// Mitsubishi GX Works2 project: 70常温静置库1130   PLC: Q10UDEH (continued)
		m_iCoordinateY:=1;
		FanucRobotIO.io_xMutexLock:=0;
	END_IF;
	IF ConveyorIO.xEmpty AND PackCommunicationIO.o_iSinglePackDonePLCPC=1 THEN
		m_iStep:=1;
	END_IF;
END_CASE;
END_FUNCTION_BLOCK

PROGRAM POU
VAR
  Conveyor70101 : Conveyor;
  Conveyor70102 : Conveyor;
  Conveyor70103 : Conveyor;
  Conveyor70104 : Conveyor;
  Conveyor70105 : Conveyor;
  Conveyor70106 : Conveyor;
  Conveyor70107 : Conveyor;
  Conveyor70108 : Conveyor;
  Conveyor70109 : Conveyor;
  Conveyor70110 : Conveyor;
  Conveyor70111 : Conveyor;
  Conveyor70112 : Conveyor;
  Conveyor70113 : Conveyor;
  Conveyor70114 : Conveyor;
  Conveyor70115 : Conveyor;
  Conveyor70116 : Conveyor;
  Conveyor70117 : Conveyor;
  Conveyor70118 : Conveyor;
  Conveyor70119 : Conveyor;
  Conveyor70120 : Conveyor;
  Conveyor70121 : Conveyor;
  Conveyor70122 : Conveyor;
  Conveyor70123 : Conveyor;
  Conveyor70124 : Conveyor;
  Conveyor70125 : Conveyor;
  Conveyor70126 : Conveyor;
  Conveyor70127 : Conveyor;
  Conveyor70128 : Conveyor;
  Conveyor70129 : Conveyor;
  Conveyor70130 : Conveyor;
  Conveyor70131 : Conveyor;
  Conveyor70132 : Conveyor;
  Conveyor70133 : Conveyor;
  Conveyor70134 : Conveyor;
  Conveyor70135 : Conveyor;
  Conveyor70136 : Conveyor;
  Conveyor70137 : Conveyor;
  Conveyor70138 : Conveyor;
  Conveyor70139 : Conveyor;
  Conveyor70140 : Conveyor;
  Conveyor70141 : Conveyor;
  Conveyor70142 : Conveyor;
  Conveyor70143 : Conveyor;
  Conveyor70144 : Conveyor;
  Conveyor70145 : Conveyor;
  Conveyor70146 : Conveyor;
  Conveyor70147 : Conveyor;
  Conveyor70148 : Conveyor;
  Conveyor70149 : Conveyor;
  Conveyor70150 : Conveyor;
  Conveyor70151 : Conveyor;
  Conveyor70152 : Conveyor;
  Conveyor70153 : Conveyor;
  Conveyor70154 : Conveyor;
  Conveyor70155 : Conveyor;
  Conveyor70156 : Conveyor;
  Conveyor70157 : Conveyor;
  Conveyor70158 : Conveyor;
  Conveyor70159 : Conveyor;
  Conveyor70160 : Conveyor;
  Conveyor70161 : Conveyor;
  Conveyor70162 : Conveyor;
  Conveyor70163 : Conveyor;
  Conveyor70164 : Conveyor;
  Conveyor70165 : Conveyor;
  Conveyor70166 : Conveyor;
  Conveyor70167 : Conveyor;
  Conveyor70168 : Conveyor;
  Conveyor70169 : Conveyor;
  Conveyor70170 : Conveyor;
  Conveyor70171 : Conveyor;
  Conveyor70172 : Conveyor;
  Conveyor70173 : Conveyor;
  Conveyor70174 : Conveyor;
  Conveyor70175 : Conveyor;
  Conveyor70176 : Conveyor;
  Conveyor70177 : Conveyor;
  Conveyor70178 : Conveyor;
  Conveyor70179 : Conveyor;
  Conveyor70180 : Conveyor;
  Conveyor70181 : Conveyor;
  Conveyor70182 : Conveyor;
  Conveyor70183 : Conveyor;
  Conveyor70184 : Conveyor;
  Conveyor70185 : Conveyor;
  Conveyor70186 : Conveyor;
  Conveyor70187 : Conveyor;
  Conveyor70188 : Conveyor;
  Conveyor70189 : Conveyor;
  Conveyor70190 : Conveyor;
  Conveyor70191 : Conveyor;
  Conveyor70192 : Conveyor;
  Conveyor70193 : Conveyor;
  Conveyor70194 : Conveyor;
  Conveyor70195 : Conveyor;
  Conveyor70196 : Conveyor;
  Conveyor70197 : Conveyor;
  Conveyor70198 : Conveyor;
  Conveyor70199 : Conveyor;
  Conveyor701100 : Conveyor;
  Conveyor701101 : Conveyor;
  Conveyor701102 : Conveyor;
  Conveyor701103 : Conveyor;
  Conveyor701104 : Conveyor;
  Conveyor701105 : Conveyor;
  Conveyor701106 : Conveyor;
  Conveyor701107 : Conveyor;
  Conveyor701108 : Conveyor;
  Conveyor701109 : Conveyor;
  Conveyor701110 : Conveyor;
  Conveyor701111 : Conveyor;
  Conveyor701112 : Conveyor;
  ConveyorIO70101 : ConveyorIO;
  ConveyorIO70102 : ConveyorIO;
  ConveyorIO70103 : ConveyorIO;
  ConveyorIO70104 : ConveyorIO;
  ConveyorIO70105 : ConveyorIO;
  ConveyorIO70106 : ConveyorIO;
  ConveyorIO70107 : ConveyorIO;
  ConveyorIO70108 : ConveyorIO;
  ConveyorIO70109 : ConveyorIO;
  ConveyorIO70110 : ConveyorIO;
  ConveyorIO70111 : ConveyorIO;
  ConveyorIO70112 : ConveyorIO;
  ConveyorIO70113 : ConveyorIO;
  ConveyorIO70114 : ConveyorIO;
  ConveyorIO70115 : ConveyorIO;
  ConveyorIO70116 : ConveyorIO;
  ConveyorIO70117 : ConveyorIO;
  ConveyorIO70118 : ConveyorIO;
  ConveyorIO70119 : ConveyorIO;
  ConveyorIO70120 : ConveyorIO;
  ConveyorIO70121 : ConveyorIO;
  ConveyorIO70122 : ConveyorIO;
  ConveyorIO70123 : ConveyorIO;
  ConveyorIO70124 : ConveyorIO;
  ConveyorIO70125 : ConveyorIO;
  ConveyorIO70126 : ConveyorIO;
  ConveyorIO70127 : ConveyorIO;
  ConveyorIO70128 : ConveyorIO;
  ConveyorIO70129 : ConveyorIO;
  ConveyorIO70130 : ConveyorIO;
  ConveyorIO70131 : ConveyorIO;
  ConveyorIO70132 : ConveyorIO;
  ConveyorIO70133 : ConveyorIO;
  ConveyorIO70134 : ConveyorIO;
  ConveyorIO70135 : ConveyorIO;
  ConveyorIO70136 : ConveyorIO;
  ConveyorIO70137 : ConveyorIO;
  ConveyorIO70138 : ConveyorIO;
  ConveyorIO70139 : ConveyorIO;
  ConveyorIO70140 : ConveyorIO;
  ConveyorIO70141 : ConveyorIO;
  ConveyorIO70142 : ConveyorIO;
  ConveyorIO70143 : ConveyorIO;
  ConveyorIO70144 : ConveyorIO;
  ConveyorIO70145 : ConveyorIO;
  ConveyorIO70146 : ConveyorIO;
  ConveyorIO70147 : ConveyorIO;
  ConveyorIO70148 : ConveyorIO;
  ConveyorIO70149 : ConveyorIO;
  ConveyorIO70150 : ConveyorIO;
  ConveyorIO70151 : ConveyorIO;
  ConveyorIO70152 : ConveyorIO;
  ConveyorIO70153 : ConveyorIO;
  ConveyorIO70154 : ConveyorIO;
  ConveyorIO70155 : ConveyorIO;
  ConveyorIO70156 : ConveyorIO;
  ConveyorIO70157 : ConveyorIO;
  ConveyorIO70158 : ConveyorIO;
  ConveyorIO70159 : ConveyorIO;
  ConveyorIO70160 : ConveyorIO;
  ConveyorIO70161 : ConveyorIO;
  ConveyorIO70162 : ConveyorIO;
  ConveyorIO70163 : ConveyorIO;
  ConveyorIO70164 : ConveyorIO;
  ConveyorIO70165 : ConveyorIO;
  ConveyorIO70166 : ConveyorIO;
  ConveyorIO70167 : ConveyorIO;
  ConveyorIO70168 : ConveyorIO;
  ConveyorIO70169 : ConveyorIO;
  ConveyorIO70170 : ConveyorIO;
  ConveyorIO70171 : ConveyorIO;
  ConveyorIO70172 : ConveyorIO;
  ConveyorIO70173 : ConveyorIO;
  ConveyorIO70174 : ConveyorIO;
  ConveyorIO70175 : ConveyorIO;
  ConveyorIO70176 : ConveyorIO;
  ConveyorIO70177 : ConveyorIO;
  ConveyorIO70178 : ConveyorIO;
  ConveyorIO70179 : ConveyorIO;
  ConveyorIO70180 : ConveyorIO;
  ConveyorIO70181 : ConveyorIO;
  ConveyorIO70182 : ConveyorIO;
  ConveyorIO70183 : ConveyorIO;
  ConveyorIO70184 : ConveyorIO;
  ConveyorIO70185 : ConveyorIO;
  ConveyorIO70186 : ConveyorIO;
  ConveyorIO70187 : ConveyorIO;
  ConveyorIO70188 : ConveyorIO;
  ConveyorIO70189 : ConveyorIO;
  ConveyorIO70190 : ConveyorIO;
  ConveyorIO70191 : ConveyorIO;
  ConveyorIO70192 : ConveyorIO;
  ConveyorIO70193 : ConveyorIO;
  ConveyorIO70194 : ConveyorIO;
  ConveyorIO70195 : ConveyorIO;
  ConveyorIO70196 : ConveyorIO;
  ConveyorIO70197 : ConveyorIO;
  ConveyorIO70198 : ConveyorIO;
  ConveyorIO70199 : ConveyorIO;
  ConveyorIO701100 : ConveyorIO;
  ConveyorIO701101 : ConveyorIO;
  ConveyorIO701102 : ConveyorIO;
  ConveyorIO701103 : ConveyorIO;
  ConveyorIO701104 : ConveyorIO;
  ConveyorIO701105 : ConveyorIO;
  ConveyorIO701106 : ConveyorIO;
  ConveyorIO701107 : ConveyorIO;
  ConveyorIO701108 : ConveyorIO;
  ConveyorIO701109 : ConveyorIO;
  ConveyorIO701110 : ConveyorIO;
  ConveyorIO701111 : ConveyorIO;
  ConveyorIO701112 : ConveyorIO;
  Switch70301 : Switch;
  SwitchIO70301 : SwitchIO;
  Lift70207 : ShuttleCar;
  LifterIO70207 : ShuttleCarIO;
  ConveyorIO701113 : ConveyorIO;
  ConveyorIO701114 : ConveyorIO;
  ConveyorIO701115 : ConveyorIO;
  ConveyorIO701116 : ConveyorIO;
  ConveyorIO701117 : ConveyorIO;
  ConveyorIO701118 : ConveyorIO;
  ConveyorIO701119 : ConveyorIO;
  ConveyorIO701120 : ConveyorIO;
  Conveyor701113 : Conveyor;
  Conveyor701114 : Conveyor;
  Conveyor701115 : Conveyor;
  Conveyor701116 : Conveyor;
  Conveyor701117 : Conveyor;
  Conveyor701118 : Conveyor;
  Conveyor701119 : Conveyor;
  Conveyor701120 : Conveyor;
  Switch70326 : Switch;
  SwitchIO70326 : SwitchIO;
  Conveyor701111_1 : Conveyor;
  ConveyorIO701111_1 : ConveyorIO;
  Switch70311 : Switch;
  SwitchIO70311 : SwitchIO;
  Switch70316 : Switch;
  SwitchIO70316 : SwitchIO;
  m_xRGVSemiAuto : BOOL;
  m_iRGVDestinationPos : INT;
  m_xRGVReset : BOOL;
  m_iRGVCurrentPos : INT;
  m_xRGVPositionArrive : BOOL;
  m_xRGVConveyorEmpty : BOOL;
  m_xRGVConveyorNextRun : BOOL;
  m_xRGVAlarm : BOOL;
  m_xtonConveyor70195Reset : TON;
  m_xtonConveyor70195CurTime : TIME;
  m_xtonConveyor70146Reset : TON;
  m_xtonConveyor70146CurTime : TIME;
  m_xtonConveyor701115Reset : TON;
  m_xtonConveyor701114Reset : TON;
  m_xtonConveyor701115CurTime : TIME;
  m_xtonConveyor701114CurTime : TIME;
  Switch70317 : Switch;
  SwitchIO70317 : SwitchIO;
  ConveyorIO70165_1 : ConveyorIO;
  Conveyor70165_1 : Conveyor;
  m_xOCV2_1LoadRequest : BOOL;  (* OCV2  1号机上料请求 *)
  m_xOCV2_1LoadStart : BOOL;  (* OCV2 1号机开始上料信号 *)
  m_xOCV2_1UnloadRequest : BOOL;  (* OCV2 1号机开始下料信号 *)
  m_xOCV2_2UnloadRequest : BOOL;  (* OCV2 2号机开始下料信号 *)
  Switch70318 : Switch;
  m_xOCV2_1UnloadStart : BOOL;  (* 允许下料 *)
  Switch70319 : Switch;
  SwitchIO70319 : SwitchIO;
  Switch70320 : Switch;
  SwitchIO70320 : SwitchIO;
  m_x60LoadRequest : BOOL;
  m_xOCV2_1LoadLock : BOOL;  (* OCV2上料自锁 *)
  m_xOCV2_1UnLoadLock : BOOL;  (* OCV2下料自锁 *)
  m_xOCV3_1LoadRequest : BOOL;  (* OCV3  1号机上料请求 *)
  m_xOCV3_1LoadStart : BOOL;  (* OCV3 1号机开始上料信号 *)
  m_xOCV3_1UnloadRequest : BOOL;  (* OCV3 1号机开始下料信号 *)
  m_xOCV3_1UnloadStart : BOOL;  (* OCV3  1号机下料请求 *)
  m_xOCV3_1LoadLock : BOOL;  (* OCV3——1上料自锁 *)
  m_xOCV3_1UnLoadLock : BOOL;  (* OCV3——1下料自锁 *)
  ConveyorIO70175_1 : ConveyorIO;
  Conveyor70175_1 : Conveyor;
  m_xtonConveyor70162Reset : TON;
  m_xtonConveyor70162CurTime : TIME;
  m_xtonConveyor701103Reset : TON;
  m_xtonConveyor701103CurTime : TIME;
  m_xtonConveyor70159Reset : TON;
  m_xtonConveyor70159CurTime : TIME;
  m_xtonConveyor701102Reset : TON;
  m_xtonConveyor701102CurTime : TIME;
  m_xtonConveyor70170Reset : TON;
  m_xtonConveyor70170CurTime : TIME;
  m_xtonConveyor70168Reset : TON;
  m_xtonConveyor70168CurTime : TIME;
  m_xOCV2_2LoadRequest : BOOL;  (* OCV2 2号机开始上料信号 *)
  m_xOCV2_2LoadStart : BOOL;  (* OCV2 2号机开始下料信号 *)
  m_xOCV2_2UnloadStart : BOOL;  (* OCV2 2号机开始下料信号 *)
  m_xOCV3_2LoadRequest : BOOL;  (* OCV3  2号机上料请求 *)
  m_xOCV3_2LoadStart : BOOL;  (* OCV3 2号机开始上料信号 *)
  m_xOCV3_2UnloadRequest : BOOL;  (* OCV3 2号机开始下料信号 *)
  m_xOCV3_2UnloadStart : BOOL;  (* OCV3  2号机下料请求 *)
  m_xtonConveyor70156Reset : TON;
  m_xtonConveyor70156CurTime : TIME;
  m_xOCV2_2LoadLock : BOOL;  (* OCV2_2上料自锁 *)
  m_xOCV2_2UnLoadLock : BOOL;  (* OCV2_2下料自锁 *)
  m_xChoose1LoadLock : BOOL;  (* 挑选1上料自锁 *)
  m_xChoose1UnLoadLock : BOOL;  (* 挑选1下料自锁 *)
  SwitchIO70318 : SwitchIO;
  m_xChoose1LoadRequest : BOOL;  (* 挑选1上料请求 *)
  m_xChoose1LoadStart : BOOL;  (* 挑选1上料信号 *)
  m_xChoose1UnloadRequest : BOOL;  (* 挑选1下料请求 *)
  m_xChoose1UnloadStart : BOOL;  (* 挑选1下料信号 *)
  m_xChoose2LoadRequest : BOOL;  (* 挑选2上料请求 *)
  m_xChoose2LoadStart : BOOL;  (* 挑选2上料信号 *)
  m_xChoose2UnloadRequest : BOOL;  (* 挑选2下料请求 *)
  m_xChoose2UnloadStart : BOOL;  (* 挑选2下料信号 *)
  m_xChoose2LoadLock : BOOL;  (* 挑选2上料自锁 *)
  m_xChoose2UnLoadLock : BOOL;  (* 挑选2下料自锁 *)
  m_xOCV3_2LoadLock : BOOL;  (* OCV3——2上料自锁 *)
  m_xOCV3_2UnLoadLock : BOOL;  (* OCV3——2下料自锁 *)
  m_xtonConveyor70150Reset : TON;
  m_xtonConveyor70150CurTime : TIME;
  m_xtonConveyor70197Reset : TON;
  m_xtonConveyor70197CurTime : TIME;
  m_xtonConveyor70148Reset : TON;
  m_xtonConveyor70148CurTime : TIME;
  m_xtonConveyor70154Reset : TON;
  m_xtonConveyor70154CurTime : TIME;
  m_xtonConveyor70199Reset : TON;
  m_xtonConveyor70199CurTime : TIME;
  ConveyorIO70173_1 : ConveyorIO;
  Conveyor70173_1 : Conveyor;
  Conveyor70184_1 : Conveyor;
  ConveyorIO70184_1 : ConveyorIO;
  m_xtonConveyor70175_1Reset : TON;
  m_xtonConveyor70175_1CurTime : TIME;
  m_xtonConveyor70141Reset : TON;
  m_xtonConveyor70141CurTime : TIME;
  m_xtonConveyor70181Reset : TON;
  m_xtonConveyor70181CurTime : TIME;
  m_xtonConveyor70174Reset : TON;
  m_xtonConveyor70174CurTime : TIME;
  Lift70208 : ShuttleCar;
  LifterIO70208 : ShuttleCarIO;
  ComConveyor70104 : ConveyorCommunication;
  ComConveyor70106 : ConveyorCommunication;
  ComConveyor70111 : ConveyorCommunication;
  ComConveyor70112 : ConveyorCommunication;
  ComConveyor70113 : ConveyorCommunication;
  ComConveyor70114 : ConveyorCommunication;
  ComConveyor70116 : ConveyorCommunication;
  ComConveyor70119 : ConveyorCommunication;
  ComConveyor70120 : ConveyorCommunication;
  ComConveyor70121 : ConveyorCommunication;
  ComConveyor70122 : ConveyorCommunication;
  ComConveyor70124 : ConveyorCommunication;
  ComConveyor70127 : ConveyorCommunication;
  ComConveyor70128 : ConveyorCommunication;
  ComConveyor70129 : ConveyorCommunication;
  ComConveyor70140 : ConveyorCommunication;
  ComConveyor70144 : ConveyorCommunication;
  ComConveyor70146 : ConveyorCommunication;
  ComConveyor70147 : ConveyorCommunication;
  ComConveyor70148 : ConveyorCommunication;
  ComConveyor70150 : ConveyorCommunication;
  ComConveyor70151 : ConveyorCommunication;
  ComConveyor70152 : ConveyorCommunication;
  ComConveyor70154 : ConveyorCommunication;
  ComConveyor70155 : ConveyorCommunication;
  ComConveyor70156 : ConveyorCommunication;
  ComConveyor70158 : ConveyorCommunication;
  ComConveyor70159 : ConveyorCommunication;
  ComConveyor70160 : ConveyorCommunication;
  ComConveyor70162 : ConveyorCommunication;
  ComConveyor70163 : ConveyorCommunication;
  ComConveyor70164 : ConveyorCommunication;
  ComConveyor70169 : ConveyorCommunication;
  ComConveyor70170 : ConveyorCommunication;
  ComConveyor70174 : ConveyorCommunication;
  ComConveyor70184 : ConveyorCommunication;
  ComConveyor70195 : ConveyorCommunication;
  ComConveyor70196 : ConveyorCommunication;
  ComConveyor70197 : ConveyorCommunication;
  ComConveyor70198 : ConveyorCommunication;
  ComConveyor70199 : ConveyorCommunication;
  ComConveyor70201 : ConveyorCommunication;
  ComConveyor70202 : ConveyorCommunication;
  ComConveyor70203 : ConveyorCommunication;
  ComConveyor70205 : ConveyorCommunication;
  ComConveyor70210 : ConveyorCommunication;
  ComConveyor701100 : ConveyorCommunication;
  ComConveyor701101 : ConveyorCommunication;
  ComConveyor701102 : ConveyorCommunication;
  ComConveyor701103 : ConveyorCommunication;
  ComConveyor701104 : ConveyorCommunication;
  ComConveyor701105 : ConveyorCommunication;
  ComConveyor701106 : ConveyorCommunication;
  ComConveyor701107 : ConveyorCommunication;
  ComConveyor701108 : ConveyorCommunication;
  ComConveyor701109 : ConveyorCommunication;
  ComConveyor701110 : ConveyorCommunication;
  ComConveyor701111 : ConveyorCommunication;
  ComConveyor701114 : ConveyorCommunication;
  ComConveyor701115 : ConveyorCommunication;
  ComConveyor701116 : ConveyorCommunication;
  ComConveyor701119 : ConveyorCommunication;
  ComConveyor701120 : ConveyorCommunication;
  ComConveyorIO70104 : CommunicationIO;
  ComConveyorIO70106 : CommunicationIO;
  ComConveyorIO70111 : CommunicationIO;
  ComConveyorIO70112 : CommunicationIO;
  ComConveyorIO70113 : CommunicationIO;
  ComConveyorIO70114 : CommunicationIO;
  ComConveyorIO70116 : CommunicationIO;
  ComConveyorIO70119 : CommunicationIO;
  ComConveyorIO70120 : CommunicationIO;
  ComConveyorIO70121 : CommunicationIO;
  ComConveyorIO70122 : CommunicationIO;
  ComConveyorIO70124 : CommunicationIO;
  ComConveyorIO70127 : CommunicationIO;
  ComConveyorIO70128 : CommunicationIO;
  ComConveyorIO70129 : CommunicationIO;
  ComConveyorIO70140 : CommunicationIO;
  ComConveyorIO70144 : CommunicationIO;
  ComConveyorIO70146 : CommunicationIO;
  ComConveyorIO70147 : CommunicationIO;
  ComConveyorIO70148 : CommunicationIO;
  ComConveyorIO70150 : CommunicationIO;
  ComConveyorIO70151 : CommunicationIO;
  ComConveyorIO70152 : CommunicationIO;
  ComConveyorIO70154 : CommunicationIO;
  ComConveyorIO70155 : CommunicationIO;
  ComConveyorIO70156 : CommunicationIO;
  ComConveyorIO70158 : CommunicationIO;
  ComConveyorIO70159 : CommunicationIO;
  ComConveyorIO70160 : CommunicationIO;
  ComConveyorIO70162 : CommunicationIO;
  ComConveyorIO70163 : CommunicationIO;
  ComConveyorIO70164 : CommunicationIO;
  ComConveyorIO70169 : CommunicationIO;
  ComConveyorIO70170 : CommunicationIO;
  ComConveyorIO70174 : CommunicationIO;
  ComConveyorIO70184 : CommunicationIO;
  ComConveyorIO70195 : CommunicationIO;
  ComConveyorIO70196 : CommunicationIO;
  ComConveyorIO70197 : CommunicationIO;
  ComConveyorIO70198 : CommunicationIO;
  ComConveyorIO70199 : CommunicationIO;
  ComConveyorIO701100 : CommunicationIO;
  ComConveyorIO701101 : CommunicationIO;
  ComConveyorIO701102 : CommunicationIO;
  ComConveyorIO701103 : CommunicationIO;
  ComConveyorIO701104 : CommunicationIO;
  ComConveyorIO701105 : CommunicationIO;
  ComConveyorIO701106 : CommunicationIO;
  ComConveyorIO701107 : CommunicationIO;
  ComConveyorIO701108 : CommunicationIO;
  ComConveyorIO701109 : CommunicationIO;
  ComConveyorIO701110 : CommunicationIO;
  ComConveyorIO701111 : CommunicationIO;
  ComConveyorIO701114 : CommunicationIO;
  ComConveyorIO701115 : CommunicationIO;
  ComConveyorIO701116 : CommunicationIO;
  ComConveyorIO701119 : CommunicationIO;
  ComConveyorIO701120 : CommunicationIO;
  m_xtonConveyor70196Reset : TON;
  m_xtonConveyor70147Reset : TON;
  m_xtonConveyor70196CurTime : TIME;
  m_xtonConveyor70147CurTime : TIME;
  Folder70201 : Folder;
  FolderIO70201 : FolderIO;
  m_xFolder70201Atuo : BOOL;
  Conveyor70148_1 : Conveyor;
  ConveyorIO70148_1 : ConveyorIO;
  Switch70312 : Switch;
  SwitchIO70312 : SwitchIO;
  DivideFolder70206 : DivideFolder;
  DivideFolderIO70206 : FolderIO;
  DivideFolder70204 : DivideFolder;
  DivideFolderIO70204 : FolderIO;
  m_xDivideFolder70204Auto : BOOL;
  ConveyorIO70165_2 : ConveyorIO;
  Conveyor70165_2 : Conveyor;
  m_xtonConveyor70164Reset : TON;
  m_xtonConveyor70164CurTime : TIME;
  m_xtonConveyor70165_1Reset : TON;
  m_xtonConveyor70165_1CurTime : TIME;
  Conveyor70168_1 : Conveyor;
  ConveyorIO70168_1 : ConveyorIO;
  Folder70205 : FolderII;
  FolderIO70205 : FolderIO;
  m_xFolder70205Atuo : BOOL;
  SortCommunication70210 : SortCommunication;  (* OCV2分拣通信 *)
  SortCommunicationIO70210 : SortCommunicationIO;  (* OCV2分拣通信 *)
  RobotIO70210 : FanucRobotIO;  (* OCV2分拣机器人 *)
  m_xDivideFolder70206Auto : BOOL;
  ConveyorIO70175_2 : ConveyorIO;
  Conveyor70175_2 : Conveyor;
  Conveyor70140_1 : Conveyor;
  ConveyorIO70140_1 : ConveyorIO;
  Switch70313 : Switch;
  SwitchIO70313 : SwitchIO;
  m_xtonConveyor701100Reset : TON;
  m_xtonConveyor70155Reset : TON;
  m_xtonConveyor701100CurTime : TIME;
  m_xtonConveyor70155CurTime : TIME;
  switch70315 : Switch;
  SwitchIO70315 : SwitchIO;
  m_xtonConveyor701104Reset : TON;
  m_xtonConveyor70163Reset : TON;
  m_xtonConveyor701104CurTime : TIME;
  m_xtonConveyor70163CurTime : TIME;
  m_xtonConveyor701120Reset : TON;
  m_xtonConveyor701120CurTime : TIME;
  m_xtonConveyor701119CurTime : TIME;
  m_xtonConveyor701119Reset : Ton;
  switch70327 : Switch;
  SwitchIO70327 : SwitchIO;
  ConveyorIO701116_1 : ConveyorIO;
  Conveyor701116_1 : Conveyor;
  m_Task70312 : PreemptivePriority;
  m_Task70312Condition : ARRAY [1..13] OF BOOL;
  m_iTask70312 : INT;
  m_xtonConveyor70151Reset : TON;
  m_xtonConveyor70198Reset : TON;
  m_xtonConveyor70151CurTime : TIME;
  m_xtonConveyor70198CurTime : TIME;
  m_Task70314 : PreemptivePriority;
  m_Task70314Condition : ARRAY [1..13] OF BOOL;
  m_iTask70314 : INT;
  m_xtonConveyor70158Reset : TON;
  m_xtonConveyor701101Reset : TON;
  m_xtonConveyor70158CurTime : TIME;
  m_xtonConveyor701101CurTime : TIME;
  Servo1 : Servo;  (* OCV2的分拣排废线 *)
  ServoIO1 : ServoIO;  (* OCV2的分拣排废线 *)
  Servo2 : Servo;  (* OCV3的分拣排废线 *)
  ServoIO2 : ServoIO;  (* OCV3的分拣排废线 *)
  ComConveyorIO70201 : CommunicationIO;
  ComConveyorIO70205 : CommunicationIO;
  SortCommunication70184 : SortCommunication;  (* OCV3分拣通信 *)
  SortCommunicationIO70184 : SortCommunicationIO;  (* OCV3分拣通信 *)
  RobotIO70184 : FanucRobotIO;  (* OCV3分拣机器人 *)
END_VAR
Conveyor70101	(ConveyorMotor:=ConveyorIO70101);
Conveyor70102	(ConveyorMotor:=ConveyorIO70102);
Conveyor70103	(ConveyorMotor:=ConveyorIO70103);
Conveyor70104	(ConveyorMotor:=ConveyorIO70104);
Conveyor70105	(ConveyorMotor:=ConveyorIO70105);
Conveyor70106	(ConveyorMotor:=ConveyorIO70106);
Conveyor70107	(ConveyorMotor:=ConveyorIO70107);
Conveyor70108	(ConveyorMotor:=ConveyorIO70108);

(*Conveyor70109	(ConveyorMotor:=ConveyorIO70109);
Conveyor70110	(ConveyorMotor:=ConveyorIO70110);
Conveyor70111	(ConveyorMotor:=ConveyorIO70111);
Conveyor70112	(ConveyorMotor:=ConveyorIO70112);
Conveyor70113	(ConveyorMotor:=ConveyorIO70113);*)
Conveyor70114	(ConveyorMotor:=ConveyorIO70114);
Conveyor70115	(ConveyorMotor:=ConveyorIO70115);
Conveyor70116	(ConveyorMotor:=ConveyorIO70116);
(*Conveyor70117	(ConveyorMotor:=ConveyorIO70117);
Conveyor70118	(ConveyorMotor:=ConveyorIO70118);
Conveyor70119	(ConveyorMotor:=ConveyorIO70119);
Conveyor70120	(ConveyorMotor:=ConveyorIO70120);
Conveyor70121	(ConveyorMotor:=ConveyorIO70121);*)
Conveyor70122	(ConveyorMotor:=ConveyorIO70122);
Conveyor70123	(ConveyorMotor:=ConveyorIO70123);
Conveyor70124	(ConveyorMotor:=ConveyorIO70124);
(*Conveyor70125	(ConveyorMotor:=ConveyorIO70125);
Conveyor70126	(ConveyorMotor:=ConveyorIO70126);
Conveyor70127	(ConveyorMotor:=ConveyorIO70127);
Conveyor70128	(ConveyorMotor:=ConveyorIO70128);
Conveyor70129	(ConveyorMotor:=ConveyorIO70129);*)
Conveyor70130	(ConveyorMotor:=ConveyorIO70130);
Conveyor70131	(ConveyorMotor:=ConveyorIO70131);
Conveyor70132	(ConveyorMotor:=ConveyorIO70132);
Conveyor70133	(ConveyorMotor:=ConveyorIO70133);
Conveyor70134	(ConveyorMotor:=ConveyorIO70134);
Conveyor70135	(ConveyorMotor:=ConveyorIO70135);
Conveyor70136	(ConveyorMotor:=ConveyorIO70136);
Conveyor70137	(ConveyorMotor:=ConveyorIO70137);
Conveyor70138	(ConveyorMotor:=ConveyorIO70138);
Conveyor70139	(ConveyorMotor:=ConveyorIO70139);
Conveyor70140	(ConveyorMotor:=ConveyorIO70140);
Conveyor70140_1	(ConveyorMotor:=ConveyorIO70140_1);
Conveyor70141	(ConveyorMotor:=ConveyorIO70141);
Conveyor70142	(ConveyorMotor:=ConveyorIO70142);
Conveyor70143	(ConveyorMotor:=ConveyorIO70143);
Conveyor70144	(ConveyorMotor:=ConveyorIO70144);
Conveyor70145	(ConveyorMotor:=ConveyorIO70145);
Conveyor70146	(ConveyorMotor:=ConveyorIO70146);
Conveyor70147	(ConveyorMotor:=ConveyorIO70147);
Conveyor70148	(ConveyorMotor:=ConveyorIO70148);
Conveyor70148_1(ConveyorMotor:= ConveyorIO70148_1 );
Conveyor70149	(ConveyorMotor:=ConveyorIO70149);
Conveyor70150	(ConveyorMotor:=ConveyorIO70150);
Conveyor70151	(ConveyorMotor:=ConveyorIO70151);
Conveyor70152	(ConveyorMotor:=ConveyorIO70152);
Conveyor70153	(ConveyorMotor:=ConveyorIO70153);
Conveyor70154	(ConveyorMotor:=ConveyorIO70154);
Conveyor70155	(ConveyorMotor:=ConveyorIO70155);
Conveyor70156	(ConveyorMotor:=ConveyorIO70156);
Conveyor70157	(ConveyorMotor:=ConveyorIO70157);
Conveyor70158	(ConveyorMotor:=ConveyorIO70158);
Conveyor70159	(ConveyorMotor:=ConveyorIO70159);
Conveyor70160	(ConveyorMotor:=ConveyorIO70160);
Conveyor70161	(ConveyorMotor:=ConveyorIO70161);
Conveyor70162	(ConveyorMotor:=ConveyorIO70162);
Conveyor70163	(ConveyorMotor:=ConveyorIO70163);
Conveyor70164	(ConveyorMotor:=ConveyorIO70164);
Conveyor70165	(ConveyorMotor:=ConveyorIO70165);
Conveyor70165_1(ConveyorMotor:= ConveyorIO70165_1 );
Conveyor70165_2(ConveyorMotor:= ConveyorIO70165_2 );
Conveyor70166	(ConveyorMotor:=ConveyorIO70166);
Conveyor70167	(ConveyorMotor:=ConveyorIO70167);
Conveyor70168	(ConveyorMotor:=ConveyorIO70168);
Conveyor70168_1	(ConveyorMotor:=ConveyorIO70168_1);
Conveyor70169	(ConveyorMotor:=ConveyorIO70169);
Conveyor70170	(ConveyorMotor:=ConveyorIO70170);
Conveyor70171	(ConveyorMotor:=ConveyorIO70171);
Conveyor70172	(ConveyorMotor:=ConveyorIO70172);
Conveyor70173	(ConveyorMotor:=ConveyorIO70173);
Conveyor70173_1	(ConveyorMotor:=ConveyorIO70173_1);
Conveyor70174	(ConveyorMotor:=ConveyorIO70174);
Conveyor70175	(ConveyorMotor:=ConveyorIO70175);
Conveyor70175_1	(ConveyorMotor:=ConveyorIO70175_1);
Conveyor70175_2	(ConveyorMotor:=ConveyorIO70175_2);
Conveyor70176	(ConveyorMotor:=ConveyorIO70176);
Conveyor70177	(ConveyorMotor:=ConveyorIO70177);
Conveyor70178	(ConveyorMotor:=ConveyorIO70178);
Conveyor70179	(ConveyorMotor:=ConveyorIO70179);
Conveyor70180	(ConveyorMotor:=ConveyorIO70180);
Conveyor70181	(ConveyorMotor:=ConveyorIO70181);
Conveyor70182	(ConveyorMotor:=ConveyorIO70182);
Conveyor70183	(ConveyorMotor:=ConveyorIO70183);
Conveyor70184	(ConveyorMotor:=ConveyorIO70184);
Conveyor70184_1	(ConveyorMotor:=ConveyorIO70184_1);
Conveyor70185	(ConveyorMotor:=ConveyorIO70185);
Conveyor70186	(ConveyorMotor:=ConveyorIO70186);
(*Conveyor70187	(ConveyorMotor:=ConveyorIO70187);
Conveyor70188	(ConveyorMotor:=ConveyorIO70188);
Conveyor70189	(ConveyorMotor:=ConveyorIO70189);*)
Conveyor70190	(ConveyorMotor:=ConveyorIO70190);
Conveyor70191	(ConveyorMotor:=ConveyorIO70191);
Conveyor70192	(ConveyorMotor:=ConveyorIO70192);
Conveyor70193	(ConveyorMotor:=ConveyorIO70193);
Conveyor70194	(ConveyorMotor:=ConveyorIO70194);
Conveyor70195	(ConveyorMotor:=ConveyorIO70195);
Conveyor70196	(ConveyorMotor:=ConveyorIO70196);
Conveyor70197	(ConveyorMotor:=ConveyorIO70197);
Conveyor70198	(ConveyorMotor:=ConveyorIO70198);
Conveyor70199	(ConveyorMotor:=ConveyorIO70199);
Conveyor701100	(ConveyorMotor:=ConveyorIO701100);
Conveyor701101	(ConveyorMotor:=ConveyorIO701101);
Conveyor701102	(ConveyorMotor:=ConveyorIO701102);
Conveyor701103	(ConveyorMotor:=ConveyorIO701103);
Conveyor701104	(ConveyorMotor:=ConveyorIO701104);
(*Conveyor701105	(ConveyorMotor:=ConveyorIO701105);
Conveyor701106	(ConveyorMotor:=ConveyorIO701106);
Conveyor701107	(ConveyorMotor:=ConveyorIO701107);
Conveyor701108	(ConveyorMotor:=ConveyorIO701108);
Conveyor701109	(ConveyorMotor:=ConveyorIO701109);
Conveyor701110	(ConveyorMotor:=ConveyorIO701110);*)
Conveyor701111	(ConveyorMotor:=ConveyorIO701111);
Conveyor701111_1(ConveyorMotor:= ConveyorIO701111_1);
Conveyor701112	(ConveyorMotor:=ConveyorIO701112);
Conveyor701113	(ConveyorMotor:=ConveyorIO701113);
Conveyor701114	(ConveyorMotor:=ConveyorIO701114);
Conveyor701115	(ConveyorMotor:=ConveyorIO701115);
Conveyor701116	(ConveyorMotor:=ConveyorIO701116);
Conveyor701117	(ConveyorMotor:=ConveyorIO701117);
Conveyor701118	(ConveyorMotor:=ConveyorIO701118);
Conveyor701119	(ConveyorMotor:=ConveyorIO701119);
Conveyor701120	(ConveyorMotor:=ConveyorIO701120);

ConveyorIO70101.xCWPresent:=X8;						
Y208:=ConveyorIO70101.xMotorCW;						
ConveyorIO70101.xForward:=M500;						
M301:= NOT ConveyorIO70101.xEmpty;						
M700:=ConveyorIO70101.xError;						
ConveyorIO70101.diDeviceID:=70101;						

ConveyorIO70102.xCWPresent:=X9;						
Y209:=ConveyorIO70102.xMotorCW;						
ConveyorIO70102.xForward:=M501;						
M302:= NOT ConveyorIO70102.xEmpty;						
M701:=ConveyorIO70102.xError;						
ConveyorIO70102.diDeviceID:=70102;						

ConveyorIO70103.xCWPresent:=XA;						
Y20A:=ConveyorIO70103.xMotorCW;						
ConveyorIO70103.xForward:=M502;						
M303:= NOT ConveyorIO70103.xEmpty;						
M702:=ConveyorIO70103.xError;						
ConveyorIO70103.diDeviceID:=70103;						

ConveyorIO70104.xCWPresent:=XB;						
Y20B:=ConveyorIO70104.xMotorCW;						
ConveyorIO70104.xForward:=M503;						
M304:= NOT ConveyorIO70104.xEmpty;						
M703:=ConveyorIO70104.xError;						
ConveyorIO70104.diDeviceID:=70104;		
ConveyorIO70104.tLoadDelay:=T#5s;				

ConveyorIO70105.xCWPresent:=XB;	
ConveyorIO70105.xPosLimit:=NOT X160;					
Y20C:=ConveyorIO70105.xMotorCW;						
ConveyorIO70105.xForward:=M504;						
M305:= NOT ConveyorIO70105.xEmpty;						
M704:=ConveyorIO70105.xError;						
ConveyorIO70105.diDeviceID:=70104;						
(*提升机线体*)
(*ConveyorIO70106.xPosLimit:=XF;						
ConveyorIO70106.xNegLimit:=X10;*)						
ConveyorIO70106.xCWPresent:=XE;						
ConveyorIO70106.xCCWPresent:=XF;						
(*Y20D:=ConveyorIO70106.xMotorCW;	*)
Y212:=ConveyorIO70106.xMotorCW;	
Y213:=ConveyorIO70106.xMotorCCW;					
ConveyorIO70106.xForward:=M505;	
ConveyorIO70106.xBackward:=M610;					
M306:= NOT ConveyorIO70106.xEmpty;						
M705:=ConveyorIO70106.xError;						
ConveyorIO70106.diDeviceID:=70106;		
ConveyorIo70106.xSizeDeficientDetect:=1;

ConveyorIO70107.xPosLimit:=X13;						
ConveyorIO70107.xNegLimit:=X14;						
ConveyorIO70107.xCWPresent:=X11;						
ConveyorIO70107.xCCWPresent:=X12;						
Y20E:=ConveyorIO70107.xMotorCW;						
ConveyorIO70107.xForward:=M506;						
M307:= NOT ConveyorIO70107.xEmpty;						
M706:=ConveyorIO70107.xError;						
ConveyorIO70107.diDeviceID:=70107;						

ConveyorIO70108.xCWPresent:=X15;						
Y20F:=ConveyorIO70108.xMotorCW;						
ConveyorIO70108.xForward:=M507;						
M308:= NOT ConveyorIO70108.xEmpty;						
M707:=ConveyorIO70108.xError;						
ConveyorIO70108.diDeviceID:=70108;						

ConveyorIO70109.xCWPresent:=X16;						
Y210:=ConveyorIO70109.xMotorCW;						
Y211:=ConveyorIO70109.xMotorCCW;						
ConveyorIO70109.xForward:=M508;						
ConveyorIO70109.xBackward:=M509;						
M309:= NOT ConveyorIO70109.xEmpty;						
M708:=ConveyorIO70109.xError;						
ConveyorIO70109.diDeviceID:=70109;						

ConveyorIO70110.xCWPresent:=X17;						
(*Y212:=ConveyorIO70110.xMotorCW;						
Y213:=ConveyorIO70110.xMotorCCW;	*)					
(*ConveyorIO70110.xForward:=M510;						
ConveyorIO70110.xBackward:=M511;		*)				
M310:= NOT ConveyorIO70110.xEmpty;						
M709:=ConveyorIO70110.xError;						
ConveyorIO70110.diDeviceID:=70110;						

ConveyorIO70111.xCWPresent:=X18;						
Y214:=ConveyorIO70111.xMotorCW;						
Y215:=ConveyorIO70111.xMotorCCW;						
ConveyorIO70111.xForward:=M512;						
ConveyorIO70111.xBackward:=M513;						
M311:= NOT ConveyorIO70111.xEmpty;						
M710:=ConveyorIO70111.xError;						
ConveyorIO70111.diDeviceID:=70111;						

ConveyorIO70112.xPosLimit:=X1A;						
ConveyorIO70112.xCWPresent:=X19;						
Y216:=ConveyorIO70112.xMotorCW;						
Y217:=ConveyorIO70112.xMotorCCW;						
ConveyorIO70112.xForward:=M514;						
ConveyorIO70112.xBackward:=M515;						
M312:= NOT ConveyorIO70112.xEmpty;						
M711:=ConveyorIO70112.xError;						
ConveyorIO70112.diDeviceID:=70112;						

ConveyorIO70113.xPosLimit:=X1C;						
ConveyorIO70113.xCWPresent:=X1B;						
Y218:=ConveyorIO70113.xMotorCW;						
Y219:=ConveyorIO70113.xMotorCCW;						
ConveyorIO70113.xForward:=M516;						
ConveyorIO70113.xBackward:=M517;						
M313:= NOT ConveyorIO70113.xEmpty;						
M712:=ConveyorIO70113.xError;						
ConveyorIO70113.diDeviceID:=70113;			
ConveyorIO70113.tLoadDelay:=T#5s;			

ConveyorIO70114.xCWPresent:=X1D;						
Y21A:=ConveyorIO70114.xMotorCW;						
Y21C:=ConveyorIO70114.xMotorCCW;						
ConveyorIO70114.xForward:=M518;						
ConveyorIO70114.xBackward:=M519;						
M314:= NOT ConveyorIO70114.xEmpty;						
M713:=ConveyorIO70114.xError;						
ConveyorIO70114.diDeviceID:=70114;						

ConveyorIO70115.xCWPresent:=X1E;						
Y21B:=ConveyorIO70115.xMotorCW;						
ConveyorIO70115.xForward:=M520;						
M315:= NOT ConveyorIO70115.xEmpty;						
M714:=ConveyorIO70115.xError;						
ConveyorIO70115.diDeviceID:=70115;						

ConveyorIO70116.xCWPresent:=X1F;						
Y21C:=ConveyorIO70116.xMotorCW;						
ConveyorIO70116.xForward:=M521;						
M316:= NOT ConveyorIO70116.xEmpty;						
M715:=ConveyorIO70116.xError;						
ConveyorIO70116.diDeviceID:=70116;						

ConveyorIO70117.xCWPresent:=X20;						
Y21D:=ConveyorIO70117.xMotorCW;						
Y21E:=ConveyorIO70117.xMotorCCW;						
ConveyorIO70117.xForward:=M522;						
ConveyorIO70117.xBackward:=M523;						
M317:= NOT ConveyorIO70117.xEmpty;						
M716:=ConveyorIO70117.xError;						
ConveyorIO70117.diDeviceID:=70117;						

ConveyorIO70118.xCWPresent:=X21;						
Y21F:=ConveyorIO70118.xMotorCW;						
Y220:=ConveyorIO70118.xMotorCCW;						
ConveyorIO70118.xForward:=M524;						
ConveyorIO70118.xBackward:=M525;						
M318:= NOT ConveyorIO70118.xEmpty;						
M717:=ConveyorIO70118.xError;						
ConveyorIO70118.diDeviceID:=70118;						

ConveyorIO70119.xCWPresent:=X22;						
Y221:=ConveyorIO70119.xMotorCW;						
Y222:=ConveyorIO70119.xMotorCCW;						
ConveyorIO70119.xForward:=M526;						
ConveyorIO70119.xBackward:=M527;						
M319:= NOT ConveyorIO70119.xEmpty;						
M718:=ConveyorIO70119.xError;						
ConveyorIO70119.diDeviceID:=70119;						

ConveyorIO70120.xPosLimit:=X24;						
ConveyorIO70120.xCWPresent:=X23;						
Y223:=ConveyorIO70120.xMotorCW;						
Y224:=ConveyorIO70120.xMotorCCW;						
ConveyorIO70120.xForward:=M528;						
ConveyorIO70120.xBackward:=M529;						
M320:= NOT ConveyorIO70120.xEmpty;						
M719:=ConveyorIO70120.xError;						
ConveyorIO70120.diDeviceID:=70120;						

ConveyorIO70121.xPosLimit:=X26;						
ConveyorIO70121.xCWPresent:=X25;						
Y225:=ConveyorIO70121.xMotorCW;						
Y226:=ConveyorIO70121.xMotorCCW;						
ConveyorIO70121.xForward:=M530;						
ConveyorIO70121.xBackward:=M531;						
M321:= NOT ConveyorIO70121.xEmpty;						
M720:=ConveyorIO70121.xError;						
ConveyorIO70121.diDeviceID:=70121;						

ConveyorIO70122.xCWPresent:=X27;						
Y227:=ConveyorIO70122.xMotorCW;						
ConveyorIO70122.xForward:=M532;						
M322:= NOT ConveyorIO70122.xEmpty;						
M721:=ConveyorIO70122.xError;						
ConveyorIO70122.diDeviceID:=70122;						

ConveyorIO70123.xCWPresent:=X28;						
Y228:=ConveyorIO70123.xMotorCW;						
ConveyorIO70123.xForward:=M533;						
M323:= NOT ConveyorIO70123.xEmpty;						
M722:=ConveyorIO70123.xError;						
ConveyorIO70123.diDeviceID:=70123;						

ConveyorIO70124.xCWPresent:=X29;						
Y229:=ConveyorIO70124.xMotorCW;						
ConveyorIO70124.xForward:=M534;						
M324:= NOT ConveyorIO70124.xEmpty;						
M723:=ConveyorIO70124.xError;						
ConveyorIO70124.diDeviceID:=70124;						

ConveyorIO70125.xCWPresent:=X2A;						
Y22A:=ConveyorIO70125.xMotorCW;						
Y22B:=ConveyorIO70125.xMotorCCW;						
ConveyorIO70125.xForward:=M535;						
ConveyorIO70125.xBackward:=M536;						
M325:= NOT ConveyorIO70125.xEmpty;						
M724:=ConveyorIO70125.xError;						
ConveyorIO70125.diDeviceID:=70125;						

